// TIA Portal project "TNprojINZ" (V15.1) (continued)
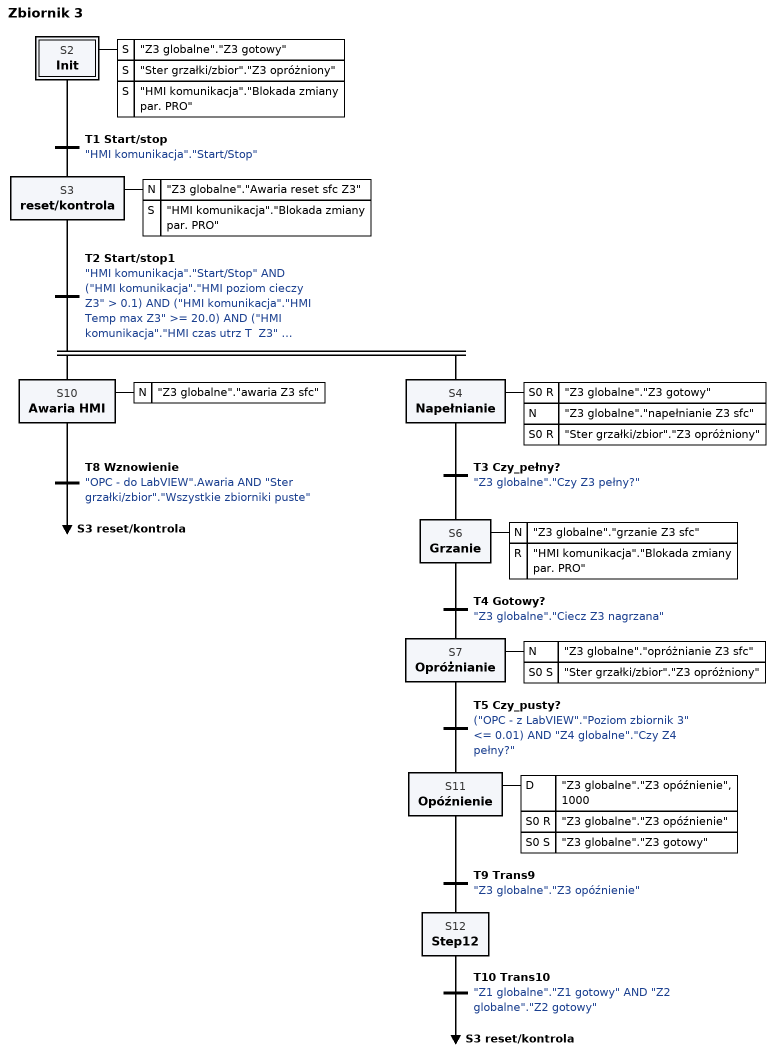
   // sequencer 1
   INITIAL_STEP Init:   // S2, max time T#10S, warning time T#7S
              S    "Z3 globalne"."Z3 gotowy"
              S    "Ster grzałki/zbior"."Z3 opróżniony"
              S    "HMI komunikacja"."Blokada zmiany par. PRO"
   END_STEP
   TRANSITION "Start/stop" FROM Init TO "reset/kontrola"   // T1
      := "HMI komunikacja"."Start/Stop";
   END_TRANSITION
   STEP "reset/kontrola":   // S3, max time T#10S, warning time T#7S
              N    "Z3 globalne"."Awaria reset sfc Z3"
              S    "HMI komunikacja"."Blokada zmiany par. PRO"
   END_STEP
   TRANSITION "Start/stop1" FROM "reset/kontrola" TO ("Awaria HMI", Napełnianie)   // T2
      := "HMI komunikacja"."Start/Stop" AND ("HMI komunikacja"."HMI poziom cieczy Z3" > 0.1) AND ("HMI komunikacja"."HMI Temp max Z3" >= 20.0) AND ("HMI komunikacja"."HMI czas utrz T  Z3" > 0.1) AND "Z1 globalne"."Z1 gotowy" AND "Z2 globalne"."Z2 gotowy";
   END_TRANSITION
   STEP Napełnianie:   // S4, max time T#10S, warning time T#7S
          S0  R    "Z3 globalne"."Z3 gotowy"
              N    "Z3 globalne"."napełnianie Z3 sfc"
          S0  R    "Ster grzałki/zbior"."Z3 opróżniony"
   END_STEP
   TRANSITION "Czy_pełny?" FROM Napełnianie TO Grzanie   // T3
      := "Z3 globalne"."Czy Z3 pełny?";
   END_TRANSITION
   STEP Grzanie:   // S6, max time T#10S, warning time T#7S
              N    "Z3 globalne"."grzanie Z3 sfc"
              R    "HMI komunikacja"."Blokada zmiany par. PRO"
   END_STEP
   TRANSITION "Gotowy?" FROM Grzanie TO Opróżnianie   // T4
      := "Z3 globalne"."Ciecz Z3 nagrzana";
   END_TRANSITION
   STEP Opróżnianie:   // S7, max time T#10S, warning time T#7S
              N    "Z3 globalne"."opróżnianie Z3 sfc"
          S0  S    "Ster grzałki/zbior"."Z3 opróżniony"
   END_STEP
   TRANSITION "Czy_pusty?" FROM Opróżnianie TO Opóźnienie   // T5
      := ("OPC - z LabVIEW"."Poziom zbiornik 3" <= 0.01) AND "Z4 globalne"."Czy Z4 pełny?";
   END_TRANSITION
   STEP "Awaria HMI":   // S10, max time T#10S, warning time T#7S
              N    "Z3 globalne"."awaria Z3 sfc"
   END_STEP
   TRANSITION Wznowienie FROM "Awaria HMI" TO "reset/kontrola"   // T8, jump
      := "OPC - do LabVIEW".Awaria AND "Ster grzałki/zbior"."Wszystkie zbiorniki puste";
   END_TRANSITION
   STEP Opóźnienie:   // S11, max time T#10S, warning time T#7S
              D    "Z3 globalne"."Z3 opóźnienie", 1000
          S0  R    "Z3 globalne"."Z3 opóźnienie"
          S0  S    "Z3 globalne"."Z3 gotowy"
   END_STEP
   TRANSITION Trans9 FROM Opóźnienie TO Step12   // T9
      := "Z3 globalne"."Z3 opóźnienie";
   END_TRANSITION
   STEP Step12:   // S12, max time T#10S, warning time T#7S
   END_STEP
   TRANSITION Trans10 FROM Step12 TO "reset/kontrola"   // T10, jump
      := "Z1 globalne"."Z1 gotowy" AND "Z2 globalne"."Z2 gotowy";
   END_TRANSITION
END_FUNCTION_BLOCK

FUNCTION_BLOCK "Zbiornik 4"   // FB4, GRAPH_PLUS
{ S7_Optimized_Access := 'TRUE' }
VERSION : 0.1
   VAR_INPUT
      OFF_SQ : Bool := false;   // Turn sequence off
      INIT_SQ : Bool := false;   // Set sequence to initial state
      ACK_EF : Bool := false;   // Acknowledge all errors and faults
      S_PREV : Bool := false;   // Output previous step in parameter S_NO
      S_NEXT : Bool := false;   // Indicate next step in parameter S_NO
      SW_AUTO : Bool := false;   // Automatic mode
      SW_TAP : Bool := false;   // Semiautomatic/switch with transition
      SW_TOP : Bool := false;   // Semiautomatic/ignore transition
      SW_MAN : Bool := false;   // Manual mode
      S_SEL : Int := 0;   // Select step to be output to S_NO
      S_ON : Bool := false;   // Activate step indicated in S_NO
      S_OFF : Bool := false;   // Deactivate step indicated S_NO
      T_PUSH : Bool := false;   // Enable transition to switch in semi automatic mode
   END_VAR
   VAR_OUTPUT
      S_NO : Int := 0;   // Step number
      S_MORE : Bool := false;   // More steps are available and can be shown in S_NO
      S_ACTIVE : Bool := false;   // Step indicated in S_NO is active
      ERR_FLT : Bool := false;   // Interlock or supervision group error
      AUTO_ON : Bool := false;   // Automatic mode is active
      TAP_ON : Bool := false;   // Semiautomatic mode/step with transition enabled
      TOP_ON : Bool := false;   // Semiautomatic mode/ignore transition enabled
      MAN_ON : Bool := false;   // Manual mode is active
   END_VAR
   VAR
      HMI_INFO : Array[0..10] of UInt;
      IF_PAR : G7_IfParPlus_V6;
      RT_DATA : G7_RTDataPlus_V6;   // Internal data area
      "Start/stop" : G7_TransitionPlus_V6;   // Transition structure
      "Start/stop1" : G7_TransitionPlus_V6;   // Transition structure
      "Czy_pełny?" : G7_TransitionPlus_V6;   // Transition structure
      "Gotowy?" : G7_TransitionPlus_V6;   // Transition structure
      "Czy_pusty?" : G7_TransitionPlus_V6;   // Transition structure
      Wznowienie : G7_TransitionPlus_V6;   // Transition structure
      Init : G7_StepPlus_V6;   // Step structure
      "reset/kontrola" : G7_StepPlus_V6;   // Step structure
      Oczekiwanie : G7_StepPlus_V6;   // Step structure
      Grzanie : G7_StepPlus_V6;   // Step structure
      Opróżnianie : G7_StepPlus_V6;   // Step structure
      "Awaria HMI" : G7_StepPlus_V6;   // Step structure
      SINI : Array[0..3] of USInt;
      LSTT : Array[0..5] of USInt;
      ATAJ : Array[0..5] of USInt;
      ATAB : Array[0..5] of USInt;
      PSTT : Array[0..5] of USInt;
      NSTT : Array[0..5] of USInt;
      ASSJ : Array[0..5] of USInt;
      ASSB : Array[0..5] of USInt;
      PTTS : Array[0..5] of USInt;
      NTTS : Array[0..5] of USInt;
      SW_SQTS : Array[0..5] of USInt;
      SWITCH : Array[0..1] of USInt;
      TVX : Array[0..3] of USInt;
      TTX : Array[0..3] of USInt;
      TSX : Array[0..3] of USInt;
      S00X : Array[0..3] of USInt;
      SOFFX : Array[0..3] of USInt;
      SONX : Array[0..3] of USInt;
      SAX : Array[0..3] of USInt;
      SERRX : Array[0..6] of USInt;
      SMX : Array[0..6] of USInt;
      S0X : Array[0..6] of USInt;
      S1X : Array[0..6] of USInt;
      IL_ALARM_INST : Diag_Alarm;
      SUP_ALARM_INST : Diag_Alarm;
      STEP_TIME_ALARM_INST : Diag_Alarm;
      IEC_TIMER_INST : IEC_TIMER;
      TRANSACTION_FLAG : Bool := false;
   END_VAR
   // SINI[0] := 2;
   // SINI[2] := 255;
   // SINI[3] := 255;
   // LSTT[0] := 255;
   // LSTT[1] := 255;
   // LSTT[2] := 255;
   // LSTT[3] := 255;
   // LSTT[4] := 1;
   // LSTT[5] := 1;
   // ATAJ[1] := 1;
   // ATAJ[2] := 2;
   // ATAJ[3] := 3;
   // ATAJ[4] := 4;
   // ATAJ[5] := 5;
   // ATAB[1] := 1;
   // ATAB[2] := 2;
   // ATAB[3] := 3;
   // ATAB[4] := 4;
   // ATAB[5] := 5;
   // PSTT[1] := 1;
   // PSTT[2] := 2;
   // PSTT[3] := 3;
   // PSTT[4] := 4;
   // PSTT[5] := 5;
   // NSTT[0] := 1;
   // NSTT[1] := 2;
   // NSTT[2] := 3;
   // NSTT[3] := 4;
   // NSTT[4] := 1;
   // NSTT[5] := 1;
   // ASSJ[1] := 1;
   // ASSJ[2] := 2;
   // ASSJ[3] := 3;
   // ASSJ[4] := 4;
   // ASSJ[5] := 5;
   // ASSB[1] := 1;
   // ASSB[2] := 5;
   // ASSB[3] := 3;
   // ASSB[4] := 4;
   // ASSB[5] := 2;
   // PTTS[0] := 255;
   // PTTS[2] := 1;
   // PTTS[3] := 2;
   // PTTS[4] := 3;
   // PTTS[5] := 1;
   // NTTS[1] := 1;
   // NTTS[2] := 2;
   // NTTS[3] := 3;
   // NTTS[4] := 4;
   // NTTS[5] := 5;
   // SW_SQTS[2] := 1;
   // SW_SQTS[3] := 1;
   // SW_SQTS[4] := 1;
   // SW_SQTS[5] := 2;
   // SWITCH[0] := 160;
   // TVX[0] := 16#1;
   // TTX[0] := 16#1;
   // TSX[0] := 16#1;
   // S00X[0] := 16#1;
   // SOFFX[0] := 16#1;
   // SONX[0] := 16#1;
   // SAX[0] := 16#1;
   // SERRX[0] := 16#1;
   // SMX[0] := 16#1;
   // S0X[0] := 16#1;
   // S1X[0] := 16#1;
BEGIN
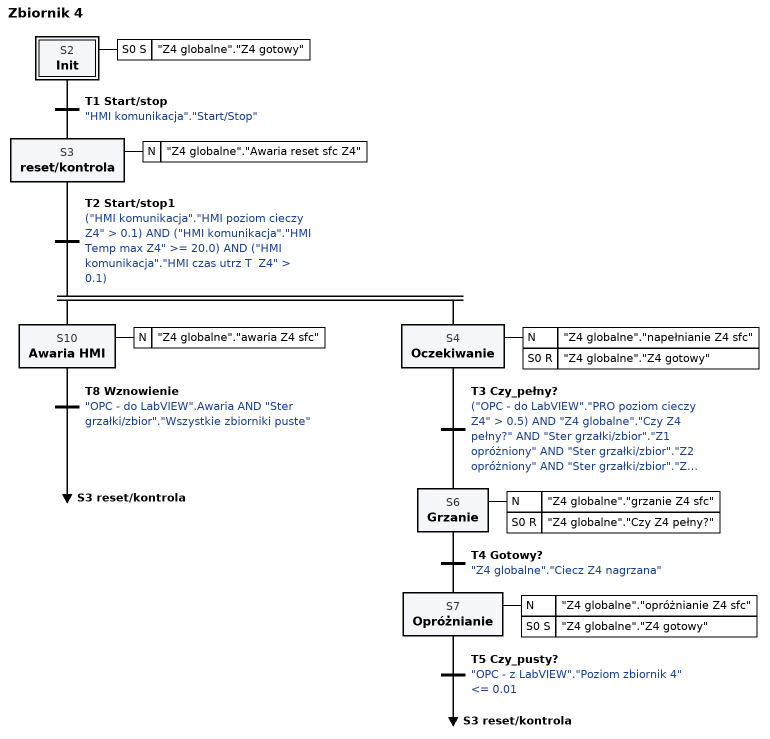
   // sequencer 1
   INITIAL_STEP Init:   // S2, max time T#10S, warning time T#7S
          S0  S    "Z4 globalne"."Z4 gotowy"
   END_STEP
   TRANSITION "Start/stop" FROM Init TO "reset/kontrola"   // T1
      := "HMI komunikacja"."Start/Stop";
   END_TRANSITION
   STEP "reset/kontrola":   // S3, max time T#10S, warning time T#7S
              N    "Z4 globalne"."Awaria reset sfc Z4"
   END_STEP
   TRANSITION "Start/stop1" FROM "reset/kontrola" TO ("Awaria HMI", Oczekiwanie)   // T2
      := ("HMI komunikacja"."HMI poziom cieczy Z4" > 0.1) AND ("HMI komunikacja"."HMI Temp max Z4" >= 20.0) AND ("HMI komunikacja"."HMI czas utrz T  Z4" > 0.1);
   END_TRANSITION
   STEP Oczekiwanie:   // S4, max time T#10S, warning time T#7S
              N    "Z4 globalne"."napełnianie Z4 sfc"
          S0  R    "Z4 globalne"."Z4 gotowy"
   END_STEP
   TRANSITION "Czy_pełny?" FROM Oczekiwanie TO Grzanie   // T3
      := ("OPC - do LabVIEW"."PRO poziom cieczy Z4" > 0.5) AND "Z4 globalne"."Czy Z4 pełny?" AND "Ster grzałki/zbior"."Z1 opróżniony" AND "Ster grzałki/zbior"."Z2 opróżniony" AND "Ster grzałki/zbior"."Z3 opróżniony";
   END_TRANSITION
   STEP Grzanie:   // S6, max time T#10S, warning time T#7S
              N    "Z4 globalne"."grzanie Z4 sfc"
          S0  R    "Z4 globalne"."Czy Z4 pełny?"
   END_STEP
   TRANSITION "Gotowy?" FROM Grzanie TO Opróżnianie   // T4
      := "Z4 globalne"."Ciecz Z4 nagrzana";
   END_TRANSITION
   STEP Opróżnianie:   // S7, max time T#10S, warning time T#7S
              N    "Z4 globalne"."opróżnianie Z4 sfc"
          S0  S    "Z4 globalne"."Z4 gotowy"
   END_STEP
   TRANSITION "Czy_pusty?" FROM Opróżnianie TO "reset/kontrola"   // T5, jump
      := "OPC - z LabVIEW"."Poziom zbiornik 4" <= 0.01;
   END_TRANSITION
   STEP "Awaria HMI":   // S10, max time T#10S, warning time T#7S
              N    "Z4 globalne"."awaria Z4 sfc"
   END_STEP
   TRANSITION Wznowienie FROM "Awaria HMI" TO "reset/kontrola"   // T8, jump
      := "OPC - do LabVIEW".Awaria AND "Ster grzałki/zbior"."Wszystkie zbiorniki puste";
   END_TRANSITION
END_FUNCTION_BLOCK

FUNCTION_BLOCK "SCL - Sterowanie pompami"   // FB5, SCL
{ S7_Optimized_Access := 'TRUE' }
VERSION : 0.1
BEGIN

   // przepompowywanie z1-3 może się zacząć, tylko gdy 'z4 gotowy' = 1    i Awaria = 0

   (* P1 i P2 *)
   IF "Z1 globalne"."opróżnianie Z1 sfc" = 1 AND "Z4 globalne"."Z4 gotowy" = 1 AND "OPC - do LabVIEW".Awaria = 0
       AND "OPC - z LabVIEW"."Poziom zbiornik 1" > 0.01 THEN

       IF "OPC - do LabVIEW"."HMI konserwacja P1" = 1 AND "OPC - do LabVIEW"."HMI konserwacja P2" = 0 THEN
           "OPC - do LabVIEW"."Pompa 2" := 1;
           "OPC - do LabVIEW"."Pompa 1" := 0;

       ELSIF "OPC - do LabVIEW"."HMI konserwacja P2" = 1 AND "OPC - do LabVIEW"."HMI konserwacja P1" = 0 THEN
           "OPC - do LabVIEW"."Pompa 1" := 1;
           "OPC - do LabVIEW"."Pompa 2" := 0;

       ELSIF "OPC - do LabVIEW"."HMI konserwacja P2" = 0 AND "OPC - do LabVIEW"."HMI konserwacja P1" = 0 THEN
           IF "Ster pompami"."przegrzana P1" = 0 AND "OPC - do LabVIEW"."Pompa 2" = 0 THEN
               "OPC - do LabVIEW"."Pompa 1" := 1;
           ELSIF "Ster pompami"."przegrzana P1" = 1 THEN
               "OPC - do LabVIEW"."Pompa 1" := 0;
               "OPC - do LabVIEW"."Pompa 2" := 1;
           ELSIF "Ster pompami"."przegrzana P2" = 1 THEN
               "OPC - do LabVIEW"."Pompa 1" := 1;
               "OPC - do LabVIEW"."Pompa 2" := 0;
           END_IF;

       END_IF;

   ELSE
       "OPC - do LabVIEW"."Pompa 1" := 0;
       "OPC - do LabVIEW"."Pompa 2" := 0;
   END_IF;


   (* P3 i P4 *)
   IF "Z2 globalne"."opróżnianie Z2 sfc" = 1 AND "Z4 globalne"."Z4 gotowy" = 1 AND "OPC - do LabVIEW".Awaria = 0
       AND "OPC - z LabVIEW"."Poziom zbiornik 2" > 0.01 THEN

       IF "OPC - do LabVIEW"."HMI konserwacja P3" = 1 AND "OPC - do LabVIEW"."HMI konserwacja P4" = 0 THEN
           "OPC - do LabVIEW"."Pompa 4" := 1;
           "OPC - do LabVIEW"."Pompa 3" := 0;

       ELSIF "OPC - do LabVIEW"."HMI konserwacja P4" = 1 AND "OPC - do LabVIEW"."HMI konserwacja P3" = 0 THEN
           "OPC - do LabVIEW"."Pompa 3" := 1;
           "OPC - do LabVIEW"."Pompa 4" := 0;

       ELSIF "OPC - do LabVIEW"."HMI konserwacja P4" = 0 AND "OPC - do LabVIEW"."HMI konserwacja P3" = 0 THEN
           IF "Ster pompami"."przegrzana P3" = 0 AND "OPC - do LabVIEW"."Pompa 4" = 0 THEN
               "OPC - do LabVIEW"."Pompa 3" := 1;
           ELSIF "Ster pompami"."przegrzana P3" = 1 THEN
               "OPC - do LabVIEW"."Pompa 3" := 0;
               "OPC - do LabVIEW"."Pompa 4" := 1;
           ELSIF "Ster pompami"."przegrzana P4" = 1 THEN
               "OPC - do LabVIEW"."Pompa 3" := 1;
               "OPC - do LabVIEW"."Pompa 4" := 0;
           END_IF;

       END_IF;

   ELSE
       "OPC - do LabVIEW"."Pompa 3" := 0;
       "OPC - do LabVIEW"."Pompa 4" := 0;
   END_IF;


   (* P5 i P6 *)
   IF "Z3 globalne"."opróżnianie Z3 sfc" = 1 AND "Z4 globalne"."Z4 gotowy" = 1 AND "OPC - do LabVIEW".Awaria = 0
       AND "OPC - z LabVIEW"."Poziom zbiornik 3" > 0.01 THEN

       IF "OPC - do LabVIEW"."HMI konserwacja P5" = 1 AND "OPC - do LabVIEW"."HMI konserwacja P6" = 0 THEN
           "OPC - do LabVIEW"."Pompa 6" := 1;
           "OPC - do LabVIEW"."Pompa 5" := 0;

       ELSIF "OPC - do LabVIEW"."HMI konserwacja P6" = 1 AND "OPC - do LabVIEW"."HMI konserwacja P5" = 0 THEN
           "OPC - do LabVIEW"."Pompa 5" := 1;
           "OPC - do LabVIEW"."Pompa 6" := 0;

       ELSIF "OPC - do LabVIEW"."HMI konserwacja P6" = 0 AND "OPC - do LabVIEW"."HMI konserwacja P5" = 0 THEN
           IF "Ster pompami"."przegrzana P5" = 0 AND "OPC - do LabVIEW"."Pompa 6" = 0 THEN
               "OPC - do LabVIEW"."Pompa 5" := 1;
           ELSIF "Ster pompami"."przegrzana P5" = 1 THEN
               "OPC - do LabVIEW"."Pompa 5" := 0;
               "OPC - do LabVIEW"."Pompa 6" := 1;
           ELSIF "Ster pompami"."przegrzana P6" = 1 THEN
               "OPC - do LabVIEW"."Pompa 5" := 1;
               "OPC - do LabVIEW"."Pompa 6" := 0;
           END_IF;

       END_IF;

   ELSE
       "OPC - do LabVIEW"."Pompa 5" := 0;
       "OPC - do LabVIEW"."Pompa 6" := 0;
   END_IF;


   (* P7 i P8 *)
   IF "Z4 globalne"."opróżnianie Z4 sfc" = 1 AND "Z4 globalne"."Z4 gotowy" = 0 AND "OPC - do LabVIEW".Awaria = 0
       AND "OPC - z LabVIEW"."Poziom zbiornik 4" > 0.01 THEN

       IF "OPC - do LabVIEW"."HMI konserwacja P7" = 1 AND "OPC - do LabVIEW"."HMI konserwacja P8" = 0 THEN
           "OPC - do LabVIEW"."Pompa 8" := 1;
           "OPC - do LabVIEW"."Pompa 7" := 0;

       ELSIF "OPC - do LabVIEW"."HMI konserwacja P8" = 1 AND "OPC - do LabVIEW"."HMI konserwacja P7" = 0 THEN
           "OPC - do LabVIEW"."Pompa 7" := 1;
           "OPC - do LabVIEW"."Pompa 8" := 0;

       ELSIF "OPC - do LabVIEW"."HMI konserwacja P8" = 0 AND "OPC - do LabVIEW"."HMI konserwacja P7" = 0 THEN
           IF "Ster pompami"."przegrzana P7" = 0 AND "OPC - do LabVIEW"."Pompa 8" = 0 THEN
               "OPC - do LabVIEW"."Pompa 7" := 1;
           ELSIF "Ster pompami"."przegrzana P7" = 1 THEN
               "OPC - do LabVIEW"."Pompa 7" := 0;
               "OPC - do LabVIEW"."Pompa 8" := 1;
           ELSIF "Ster pompami"."przegrzana P8" = 1 THEN
               "OPC - do LabVIEW"."Pompa 7" := 1;
               "OPC - do LabVIEW"."Pompa 8" := 0;
           END_IF;

       END_IF;

   ELSE
       "OPC - do LabVIEW"."Pompa 7" := 0;
       "OPC - do LabVIEW"."Pompa 8" := 0;
   END_IF;
END_FUNCTION_BLOCK

FUNCTION_BLOCK "FB - grzałki"   // FB6, FBD
{ S7_Optimized_Access := 'TRUE' }
VERSION : 0.1
   VAR_IN_OUT
      SUBrhZ1a : Real;
      SUBrhZ1b : Real;
      SUBrhZ2a : Real;
      SUBrhZ2b : Real;
      SUBrhZ3a : Real;
      SUBrhZ3b : Real;
      SUBrhZ4a : Real;
      SUBrhZ4b : Real;
      czasUTRZg1 : Real;
      czasUTRZg2 : Real;
      czasUTRZg3 : Real;
      czasUTRZg4 : Real;
      KonwTimerZ1in : Time;
      KonwTimerZ2in : Time;
      KonwTimerZ3in : Time;
      KonwTimerZ4in : Time;
      KonwTimerZ1out : Time;
      KonwTimerZ2out : Time;
      KonwTimerZ3out : Time;
      KonwTimerZ4out : Time;
      KinZ1 : Real;
      KinZ2 : Real;
      KinZ3 : Real;
      KinZ4 : Real;
      KoutZ1 : Real;
      KoutZ2 : Real;
      KoutZ3 : Real;
      KoutZ4 : Real;
   END_VAR
BEGIN

REGION Network 1: Regulator histerezowy - grzałka Z1
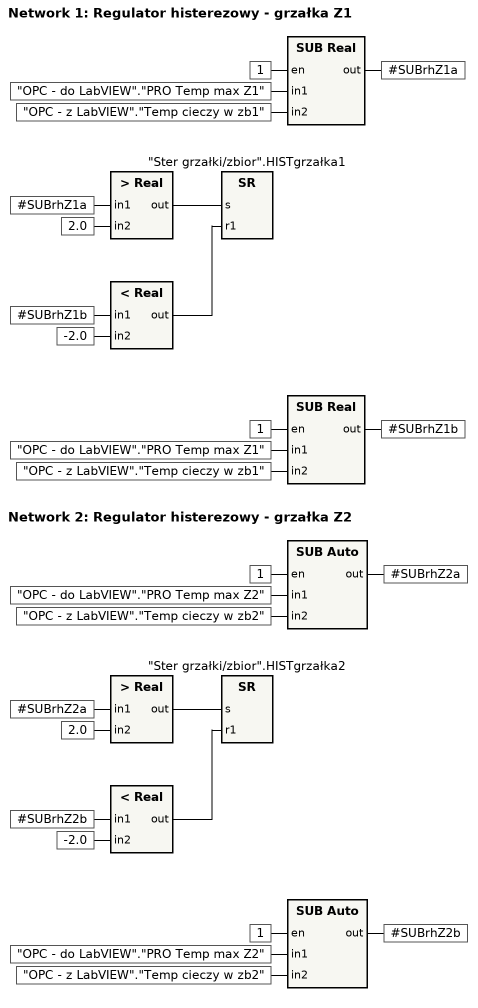
   IF 1 THEN
       #SUBrhZ1a := "OPC - do LabVIEW"."PRO Temp max Z1" - "OPC - z LabVIEW"."Temp cieczy w zb1";
   END_IF;
   IF #SUBrhZ1a > 2.0 THEN
       "Ster grzałki/zbior".HISTgrzałka1 := TRUE;   // SR flip-flop
   END_IF;
   IF #SUBrhZ1b < (-2.0) THEN "Ster grzałki/zbior".HISTgrzałka1 := FALSE; END_IF;
   IF 1 THEN
       #SUBrhZ1b := "OPC - do LabVIEW"."PRO Temp max Z1" - "OPC - z LabVIEW"."Temp cieczy w zb1";
   END_IF;
END_REGION

REGION Network 2: Regulator histerezowy - grzałka Z2
   IF 1 THEN
       #SUBrhZ2a := "OPC - do LabVIEW"."PRO Temp max Z2" - "OPC - z LabVIEW"."Temp cieczy w zb2";
   END_IF;
   IF #SUBrhZ2a > 2.0 THEN
       "Ster grzałki/zbior".HISTgrzałka2 := TRUE;   // SR flip-flop
   END_IF;
   IF #SUBrhZ2b < (-2.0) THEN "Ster grzałki/zbior".HISTgrzałka2 := FALSE; END_IF;
   IF 1 THEN
       #SUBrhZ2b := "OPC - do LabVIEW"."PRO Temp max Z2" - "OPC - z LabVIEW"."Temp cieczy w zb2";
   END_IF;
END_REGION

REGION Network 3: Regulator histerezowy - grzałka Z3
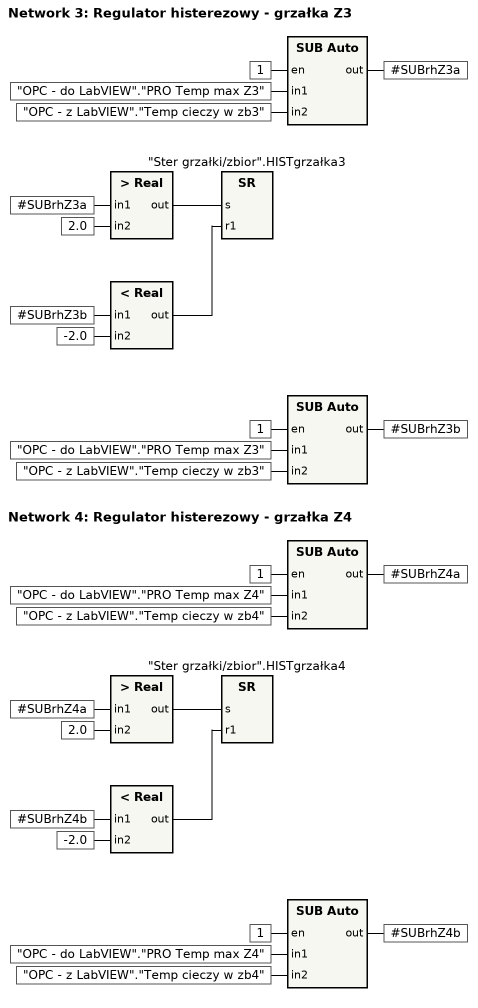
   IF 1 THEN
       #SUBrhZ3a := "OPC - do LabVIEW"."PRO Temp max Z3" - "OPC - z LabVIEW"."Temp cieczy w zb3";
   END_IF;
   IF #SUBrhZ3a > 2.0 THEN
       "Ster grzałki/zbior".HISTgrzałka3 := TRUE;   // SR flip-flop
   END_IF;
   IF #SUBrhZ3b < (-2.0) THEN "Ster grzałki/zbior".HISTgrzałka3 := FALSE; END_IF;
   IF 1 THEN
       #SUBrhZ3b := "OPC - do LabVIEW"."PRO Temp max Z3" - "OPC - z LabVIEW"."Temp cieczy w zb3";
   END_IF;
END_REGION

REGION Network 4: Regulator histerezowy - grzałka Z4
   IF 1 THEN
       #SUBrhZ4a := "OPC - do LabVIEW"."PRO Temp max Z4" - "OPC - z LabVIEW"."Temp cieczy w zb4";
   END_IF;
   IF #SUBrhZ4a > 2.0 THEN
       "Ster grzałki/zbior".HISTgrzałka4 := TRUE;   // SR flip-flop
   END_IF;
   IF #SUBrhZ4b < (-2.0) THEN "Ster grzałki/zbior".HISTgrzałka4 := FALSE; END_IF;
   IF 1 THEN
       #SUBrhZ4b := "OPC - do LabVIEW"."PRO Temp max Z4" - "OPC - z LabVIEW"."Temp cieczy w zb4";
   END_IF;
END_REGION

REGION Network 5: Czas utrzymania temp - grzałka Z1
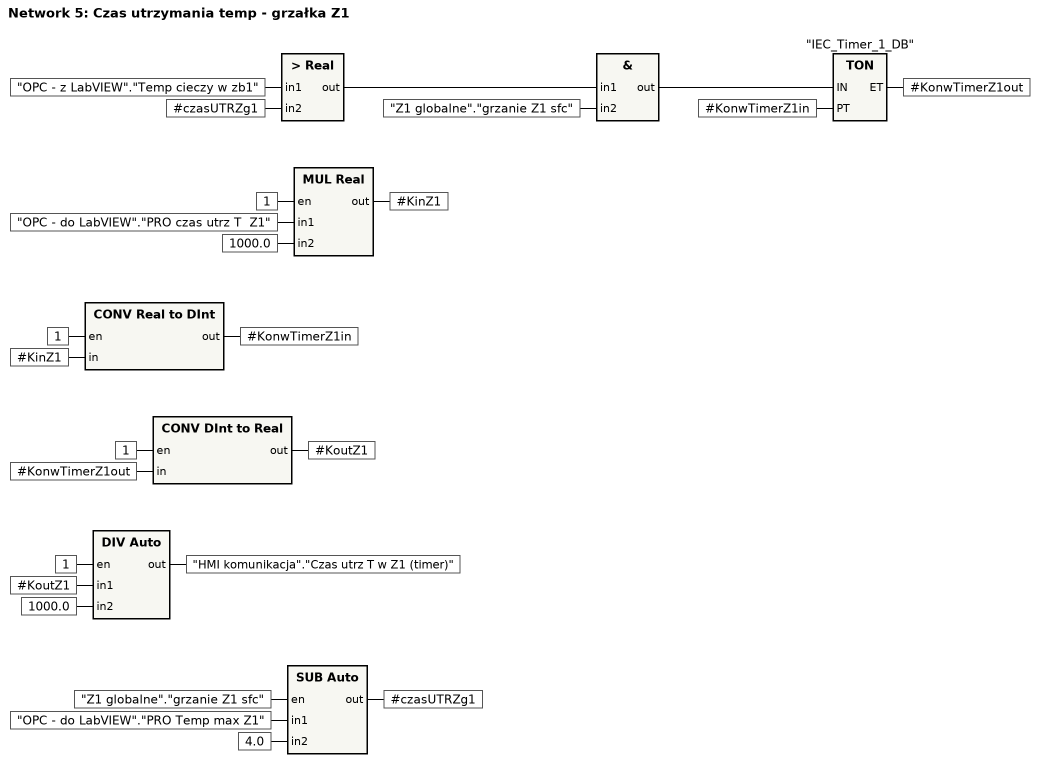
   "IEC_Timer_1_DB".TON(IN := ("OPC - z LabVIEW"."Temp cieczy w zb1" > #czasUTRZg1) AND "Z1 globalne"."grzanie Z1 sfc",
                        PT := #KonwTimerZ1in,
                        ET => #KonwTimerZ1out);
   IF 1 THEN
       #KinZ1 := "OPC - do LabVIEW"."PRO czas utrz T  Z1" * 1000.0;
       #KonwTimerZ1in := REAL_TO_DINT(#KinZ1);
       #KoutZ1 := DINT_TO_REAL(#KonwTimerZ1out);
       "HMI komunikacja"."Czas utrz T w Z1 (timer)" := #KoutZ1 / 1000.0;
   END_IF;
   IF "Z1 globalne"."grzanie Z1 sfc" THEN #czasUTRZg1 := "OPC - do LabVIEW"."PRO Temp max Z1" - 4.0; END_IF;
END_REGION

REGION Network 6: Czas utrzymania temp - grzałka Z2
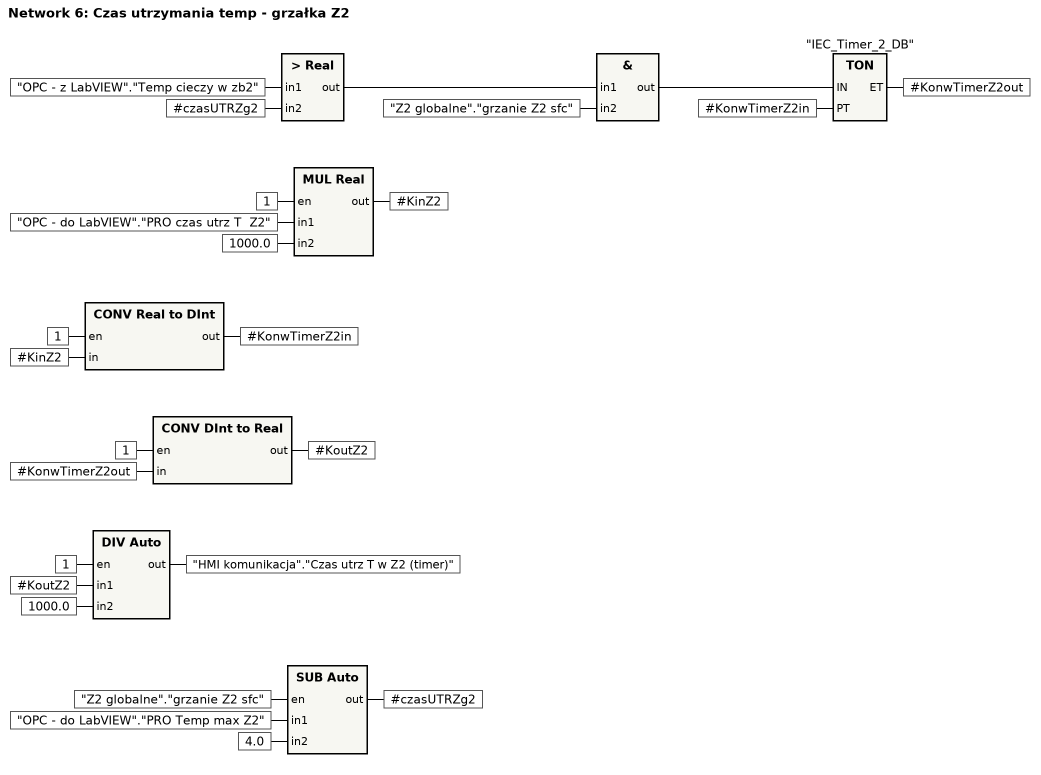
   "IEC_Timer_2_DB".TON(IN := ("OPC - z LabVIEW"."Temp cieczy w zb2" > #czasUTRZg2) AND "Z2 globalne"."grzanie Z2 sfc",
                        PT := #KonwTimerZ2in,
                        ET => #KonwTimerZ2out);
   IF 1 THEN
       #KinZ2 := "OPC - do LabVIEW"."PRO czas utrz T  Z2" * 1000.0;
       #KonwTimerZ2in := REAL_TO_DINT(#KinZ2);
       #KoutZ2 := DINT_TO_REAL(#KonwTimerZ2out);
       "HMI komunikacja"."Czas utrz T w Z2 (timer)" := #KoutZ2 / 1000.0;
   END_IF;
   IF "Z2 globalne"."grzanie Z2 sfc" THEN #czasUTRZg2 := "OPC - do LabVIEW"."PRO Temp max Z2" - 4.0; END_IF;
END_REGION

REGION Network 7: Czas utrzymania temp - grzałka Z3
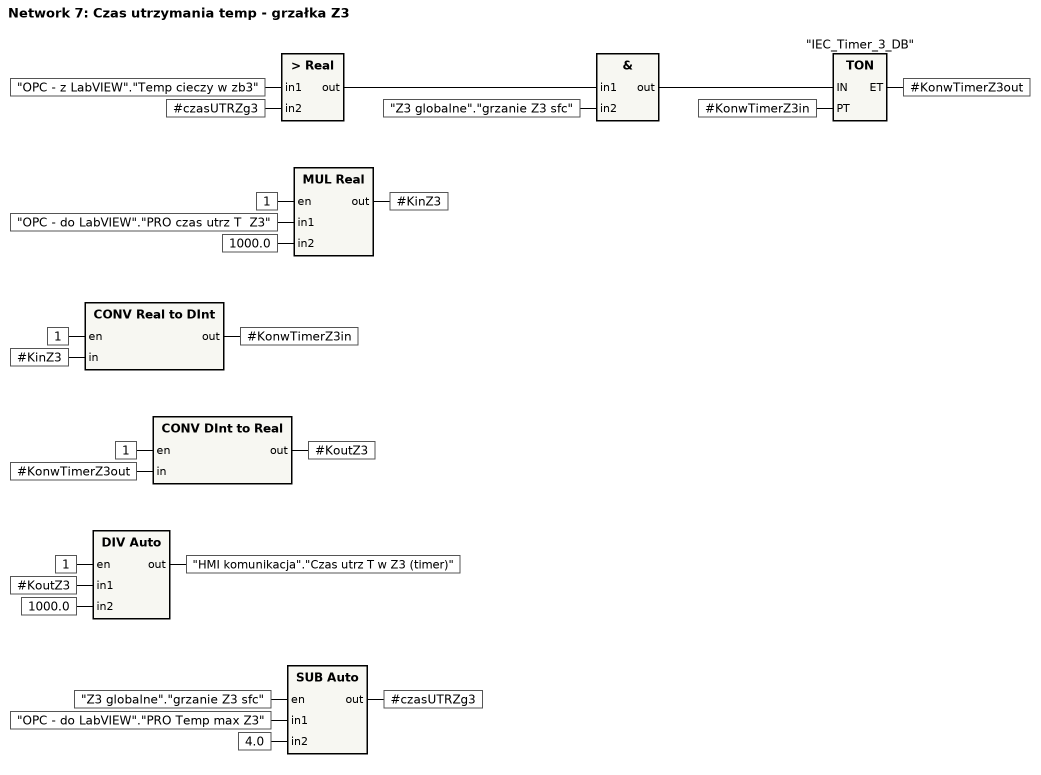
   "IEC_Timer_3_DB".TON(IN := ("OPC - z LabVIEW"."Temp cieczy w zb3" > #czasUTRZg3) AND "Z3 globalne"."grzanie Z3 sfc",
                        PT := #KonwTimerZ3in,
                        ET => #KonwTimerZ3out);
   IF 1 THEN
       #KinZ3 := "OPC - do LabVIEW"."PRO czas utrz T  Z3" * 1000.0;
       #KonwTimerZ3in := REAL_TO_DINT(#KinZ3);
       #KoutZ3 := DINT_TO_REAL(#KonwTimerZ3out);
       "HMI komunikacja"."Czas utrz T w Z3 (timer)" := #KoutZ3 / 1000.0;
   END_IF;
   IF "Z3 globalne"."grzanie Z3 sfc" THEN #czasUTRZg3 := "OPC - do LabVIEW"."PRO Temp max Z3" - 4.0; END_IF;
END_REGION

REGION Network 8: Czas utrzymania temp - grzałka Z4
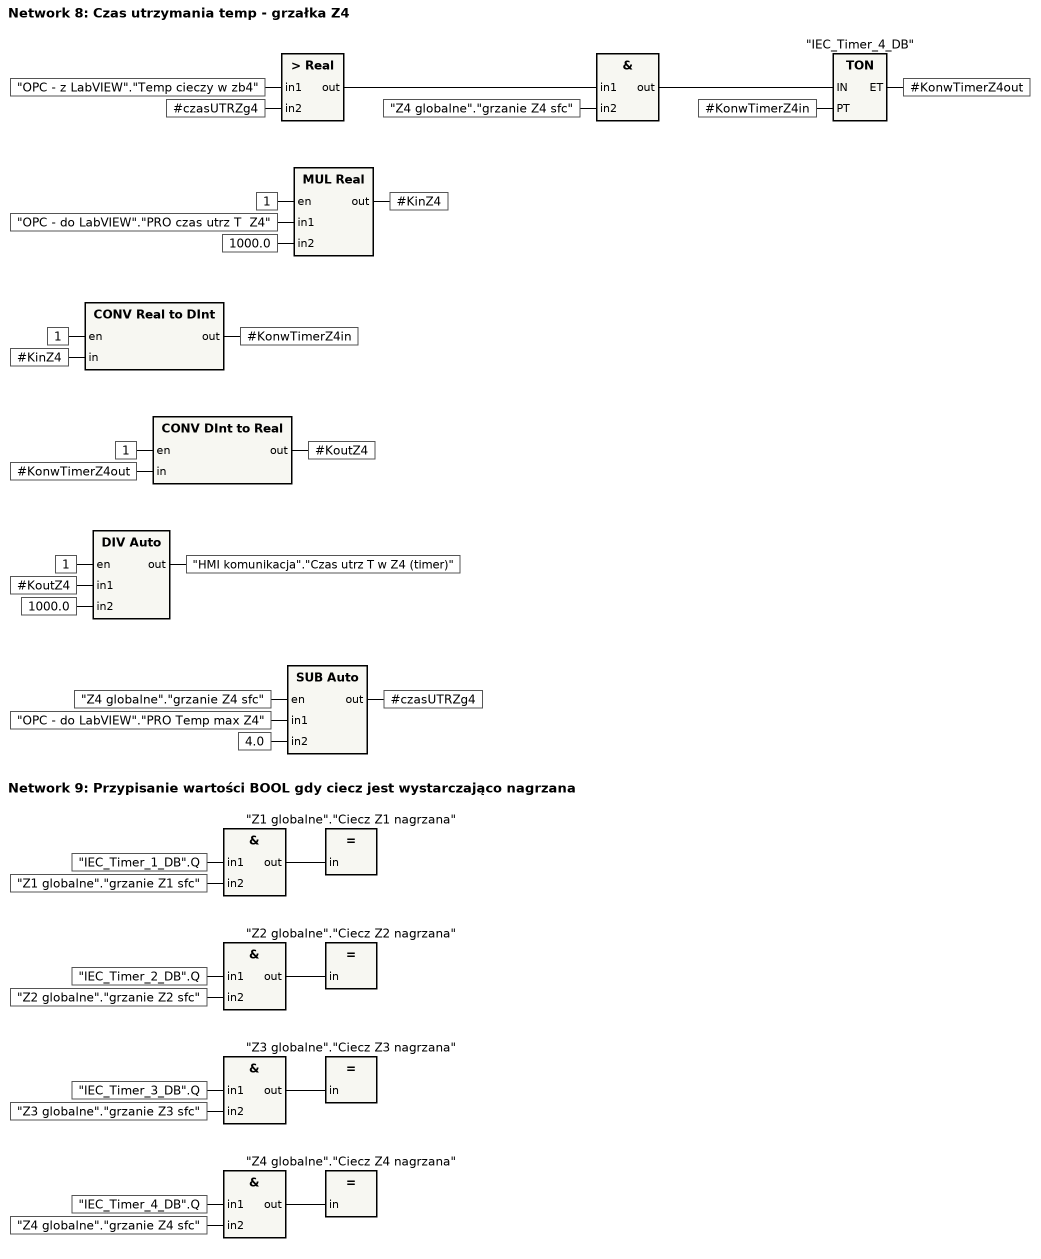
   "IEC_Timer_4_DB".TON(IN := ("OPC - z LabVIEW"."Temp cieczy w zb4" > #czasUTRZg4) AND "Z4 globalne"."grzanie Z4 sfc",
                        PT := #KonwTimerZ4in,
                        ET => #KonwTimerZ4out);
   IF 1 THEN
       #KinZ4 := "OPC - do LabVIEW"."PRO czas utrz T  Z4" * 1000.0;
       #KonwTimerZ4in := REAL_TO_DINT(#KinZ4);
       #KoutZ4 := DINT_TO_REAL(#KonwTimerZ4out);
       "HMI komunikacja"."Czas utrz T w Z4 (timer)" := #KoutZ4 / 1000.0;
   END_IF;
   IF "Z4 globalne"."grzanie Z4 sfc" THEN #czasUTRZg4 := "OPC - do LabVIEW"."PRO Temp max Z4" - 4.0; END_IF;
END_REGION

REGION Network 9: Przypisanie wartości BOOL gdy ciecz jest wystarczająco nagrzana
   "Z1 globalne"."Ciecz Z1 nagrzana" := "IEC_Timer_1_DB".Q AND "Z1 globalne"."grzanie Z1 sfc";
   "Z2 globalne"."Ciecz Z2 nagrzana" := "IEC_Timer_2_DB".Q AND "Z2 globalne"."grzanie Z2 sfc";
   "Z3 globalne"."Ciecz Z3 nagrzana" := "IEC_Timer_3_DB".Q AND "Z3 globalne"."grzanie Z3 sfc";
   "Z4 globalne"."Ciecz Z4 nagrzana" := "IEC_Timer_4_DB".Q AND "Z4 globalne"."grzanie Z4 sfc";
END_REGION
END_FUNCTION_BLOCK

FUNCTION_BLOCK "SCL - Napełnianie i kontrola"   // FB7, SCL
{ S7_Optimized_Access := 'TRUE' }
VERSION : 0.1
BEGIN
   (*
   napełnianie z1-3 zaczyna się gdy 'sfc napełnianie ... = 1'   i awaria = 0     
   pro z... = poz z HMI, gdy napełnianie z sfc = 1 - przypisanie parametru z hmi do początku procesu napeł sfc
   Pro poz z4 = pro z1 + pro z2 + pro z3  -  ok
   i inne pro = hmi również
   otwieramy zawory wlotowe
   sprawdzenie czy rzeczywisty poz z LabVIEW = (zrobić zakres +/- 1) Pro poz z... - zmienna ''czy pełny?'' w tranzycji po step napełnianie

   *)

   //Przypisanie parametrów i napełnianie Z1
   IF "Z1 globalne"."napełnianie Z1 sfc" = 1 AND "OPC - do LabVIEW".Awaria = 0 THEN
       "OPC - do LabVIEW"."PRO poziom cieczy Z1" := "HMI komunikacja"."HMI poziom cieczy Z1";
       "OPC - do LabVIEW"."PRO Temp max Z1" := "HMI komunikacja"."HMI Temp max Z1";
       "OPC - do LabVIEW"."PRO czas utrz T  Z1" := "HMI komunikacja"."HMI czas utrz T  Z1";

       //Napełnianie Z1
       IF "OPC - do LabVIEW"."PRO poziom cieczy Z1" > 15 THEN

           IF ("OPC - z LabVIEW"."Poziom zbiornik 1" > ("OPC - do LabVIEW"."PRO poziom cieczy Z1" + 1)) THEN
               "OPC - do LabVIEW"."Zawór spustowy Z1" := 1;
               "OPC - do LabVIEW"."Zawór wlotowy 1" := 0;
               "Z1 globalne"."Czy Z1 pełny?" := 0;

           ELSIF ("OPC - z LabVIEW"."Poziom zbiornik 1" >= ("OPC - do LabVIEW"."PRO poziom cieczy Z1" - 1)) AND
               ("OPC - z LabVIEW"."Poziom zbiornik 1" <= ("OPC - do LabVIEW"."PRO poziom cieczy Z1" + 1)) THEN
               "Z1 globalne"."Czy Z1 pełny?" := 1;
               "OPC - do LabVIEW"."Zawór spustowy Z1" := 0;
               "OPC - do LabVIEW"."Zawór wlotowy 1" := 0;

           ELSIF ("OPC - z LabVIEW"."Poziom zbiornik 1" < ("OPC - do LabVIEW"."PRO poziom cieczy Z1" - 1)) THEN
               "OPC - do LabVIEW"."Zawór spustowy Z1" := 0;
               "OPC - do LabVIEW"."Zawór wlotowy 1" := 1;
               "Z1 globalne"."Czy Z1 pełny?" := 0;
           END_IF;
       ELSE
           IF "OPC - z LabVIEW"."Poziom zbiornik 1" > 0.01 THEN
               "OPC - do LabVIEW"."Zawór spustowy Z1" := 1;
           ELSIF "OPC - z LabVIEW"."Poziom zbiornik 1" < 0.01 THEN
               "OPC - do LabVIEW"."Zawór spustowy Z1" := 0;
               "Z1 globalne"."Czy Z1 pełny?" := 1;
           END_IF;

       END_IF;
   ELSE
       "OPC - do LabVIEW"."Zawór wlotowy 1" := 0;
       "Z1 globalne"."Czy Z1 pełny?" := 0;
   END_IF;

   //Przypisanie parametrów i napełnianie Z2
   IF "Z2 globalne"."napełnianie Z2 sfc" = 1 AND "OPC - do LabVIEW".Awaria = 0 THEN
       "OPC - do LabVIEW"."PRO poziom cieczy Z2" := "HMI komunikacja"."HMI poziom cieczy Z2";
       "OPC - do LabVIEW"."PRO Temp max Z2" := "HMI komunikacja"."HMI Temp max Z2";
       "OPC - do LabVIEW"."PRO czas utrz T  Z2" := "HMI komunikacja"."HMI czas utrz T  Z2";

       //Napełnianie Z2
       IF "OPC - do LabVIEW"."PRO poziom cieczy Z2" > 15 THEN

           IF ("OPC - z LabVIEW"."Poziom zbiornik 2" > ("OPC - do LabVIEW"."PRO poziom cieczy Z2" + 1)) THEN
               "OPC - do LabVIEW"."Zawór spustowy Z2" := 1;
               "OPC - do LabVIEW"."Zawór wlotowy 2" := 0;
               "Z2 globalne"."Czy Z2 pełny?" := 0;

           ELSIF ("OPC - z LabVIEW"."Poziom zbiornik 2" >= ("OPC - do LabVIEW"."PRO poziom cieczy Z2" - 1)) AND
               ("OPC - z LabVIEW"."Poziom zbiornik 2" <= ("OPC - do LabVIEW"."PRO poziom cieczy Z2" + 1)) THEN
               "Z2 globalne"."Czy Z2 pełny?" := 1;
               "OPC - do LabVIEW"."Zawór spustowy Z2" := 0;
               "OPC - do LabVIEW"."Zawór wlotowy 2" := 0;

           ELSIF ("OPC - z LabVIEW"."Poziom zbiornik 2" < ("OPC - do LabVIEW"."PRO poziom cieczy Z2" - 1)) THEN
               "OPC - do LabVIEW"."Zawór spustowy Z2" := 0;
               "OPC - do LabVIEW"."Zawór wlotowy 2" := 1;
               "Z2 globalne"."Czy Z2 pełny?" := 0;
           END_IF;
       ELSE
           IF "OPC - z LabVIEW"."Poziom zbiornik 2" > 0.01 THEN
               "OPC - do LabVIEW"."Zawór spustowy Z2" := 1;
           ELSIF "OPC - z LabVIEW"."Poziom zbiornik 2" < 0.01 THEN
               "OPC - do LabVIEW"."Zawór spustowy Z2" := 0;
               "Z2 globalne"."Czy Z2 pełny?" := 1;
           END_IF;
       END_IF;
   ELSE
       "OPC - do LabVIEW"."Zawór wlotowy 2" := 0;
       "Z2 globalne"."Czy Z2 pełny?" := 0;
   END_IF;

   //Przypisanie parametrów i napełnianie Z3
   IF "Z3 globalne"."napełnianie Z3 sfc" = 1 AND "OPC - do LabVIEW".Awaria = 0 THEN
       "OPC - do LabVIEW"."PRO poziom cieczy Z3" := "HMI komunikacja"."HMI poziom cieczy Z3";
       "OPC - do LabVIEW"."PRO Temp max Z3" := "HMI komunikacja"."HMI Temp max Z3";
       "OPC - do LabVIEW"."PRO czas utrz T  Z3" := "HMI komunikacja"."HMI czas utrz T  Z3";

       //Napełnianie Z3
       IF "OPC - do LabVIEW"."PRO poziom cieczy Z3" > 15 THEN

        IF ("OPC - z LabVIEW"."Poziom zbiornik 3" > ("OPC - do LabVIEW"."PRO poziom cieczy Z3" + 1)) THEN
           "OPC - do LabVIEW"."Zawór spustowy Z3" := 1;
           "OPC - do LabVIEW"."Zawór wlotowy 3" := 0;
           "Z3 globalne"."Czy Z3 pełny?" := 0;

         ELSIF ("OPC - z LabVIEW"."Poziom zbiornik 3" >= ("OPC - do LabVIEW"."PRO poziom cieczy Z3" - 1)) AND
           ("OPC - z LabVIEW"."Poziom zbiornik 3" <= ("OPC - do LabVIEW"."PRO poziom cieczy Z3" + 1)) THEN
           "Z3 globalne"."Czy Z3 pełny?" := 1;
           "OPC - do LabVIEW"."Zawór spustowy Z3" := 0;
           "OPC - do LabVIEW"."Zawór wlotowy 3" := 0;

         ELSIF ("OPC - z LabVIEW"."Poziom zbiornik 3" < ("OPC - do LabVIEW"."PRO poziom cieczy Z3" - 1)) THEN
           "OPC - do LabVIEW"."Zawór spustowy Z3" := 0;
           "OPC - do LabVIEW"."Zawór wlotowy 3" := 1;
           "Z3 globalne"."Czy Z3 pełny?" := 0;
         END_IF;
       ELSE
           IF "OPC - z LabVIEW"."Poziom zbiornik 3" > 0.01 THEN
               "OPC - do LabVIEW"."Zawór spustowy Z3" := 1;
           ELSIF "OPC - z LabVIEW"."Poziom zbiornik 3" < 0.01 THEN
               "OPC - do LabVIEW"."Zawór spustowy Z3" := 0;
               "Z3 globalne"."Czy Z3 pełny?" := 1;
           END_IF;
       END_IF;
   ELSE
       "OPC - do LabVIEW"."Zawór wlotowy 3" := 0;
       "Z3 globalne"."Czy Z3 pełny?" := 0;
   END_IF;

   //Przypisanie parametrów i napełnianie Z4
   IF "Z4 globalne"."napełnianie Z4 sfc" = 1 AND "OPC - do LabVIEW".Awaria = 0 THEN
       "OPC - do LabVIEW"."PRO poziom cieczy Z4" := "OPC - do LabVIEW"."PRO poziom cieczy Z1" + "OPC - do LabVIEW"."PRO poziom cieczy Z2" + "OPC - do LabVIEW"."PRO poziom cieczy Z3";
       "OPC - do LabVIEW"."PRO Temp max Z4" := "HMI komunikacja"."HMI Temp max Z4";
       "OPC - do LabVIEW"."PRO czas utrz T  Z4" := "HMI komunikacja"."HMI czas utrz T  Z4";

       //Napełnianie Z1
       IF ("OPC - z LabVIEW"."Poziom zbiornik 4" >= ("OPC - do LabVIEW"."PRO poziom cieczy Z4" - 3)) AND
           ("OPC - z LabVIEW"."Poziom zbiornik 4" <= ("OPC - do LabVIEW"."PRO poziom cieczy Z4" + 3)) THEN
           //AND
           //"Ster grzałki/zbior"."Z1 opróżniony" = 1 AND "Ster grzałki/zbior"."Z2 opróżniony" = 1 AND "Ster grzałki/zbior"."Z3 opróżniony" = 1
           "Z4 globalne"."Czy Z4 pełny?" := 1;
           "OPC - do LabVIEW"."Zawór spustowy Z4" := 0;